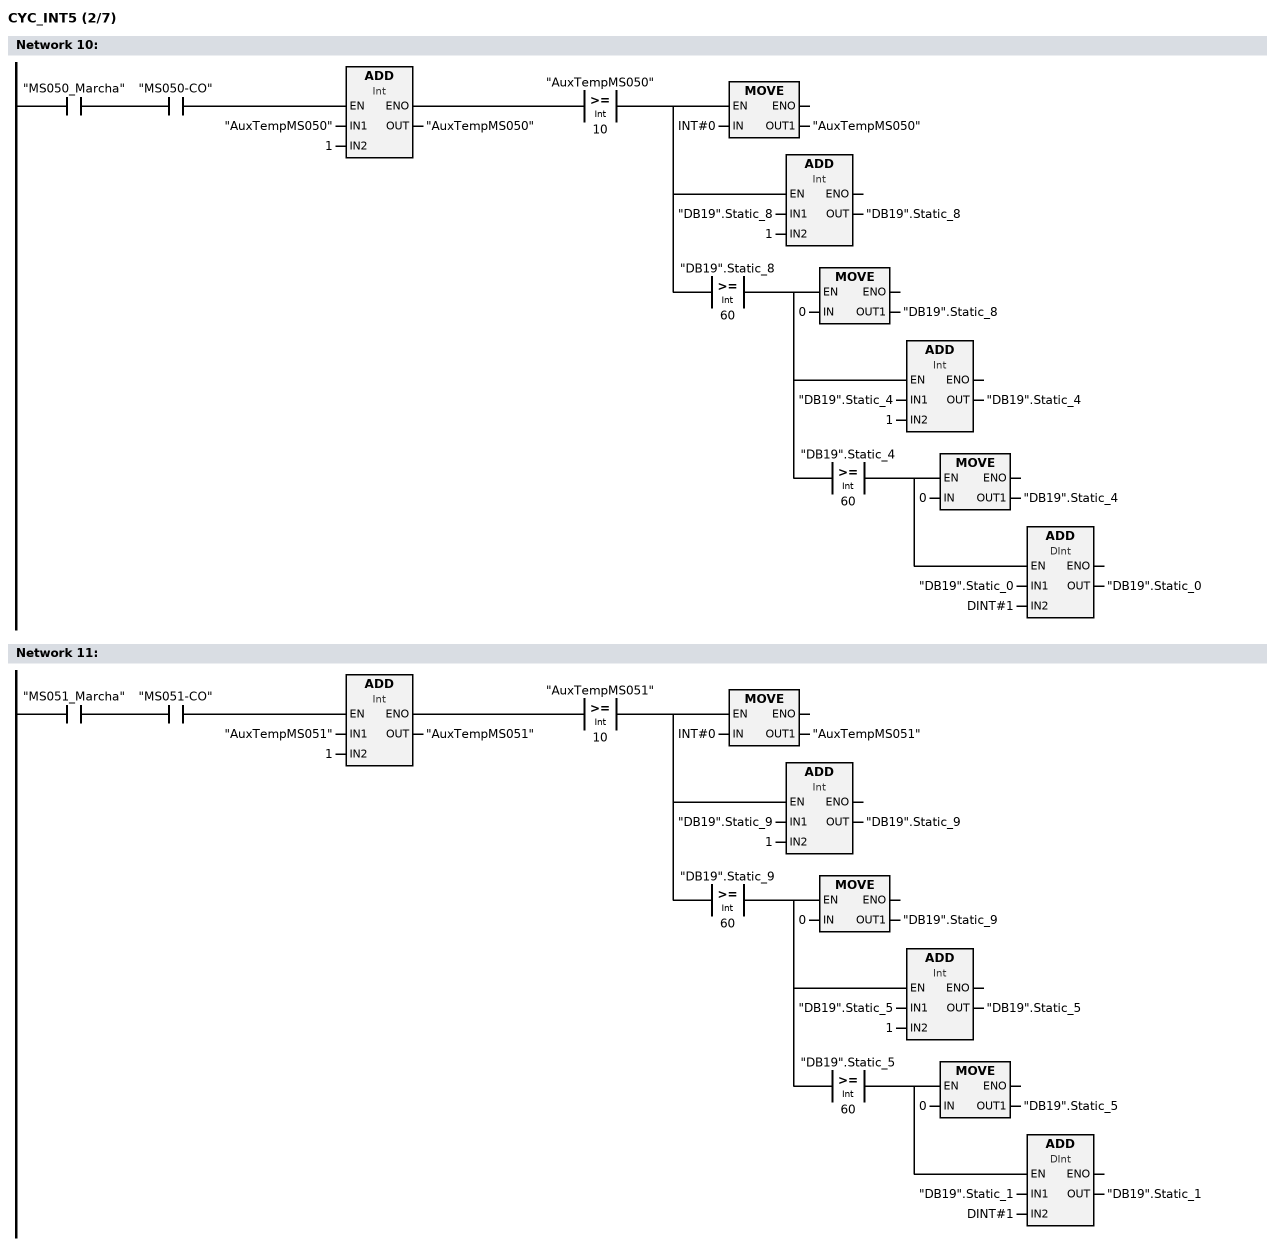
   RUNG wire#powerrail
      Contact( "MS050_Marcha" )
      Contact( "MS050-CO" )
      { S7_Templates := "SrcType := Int"; S7_GenerateENO := "TRUE" } Add(in1 := "AuxTempMS050", in2 := 1, out => "AuxTempMS050")
      { S7_Templates := "SrcType := Int" } GE_Contact(in1 := "AuxTempMS050", in2 := 10)
      wire#w1
      { S7_GenerateENO := "TRUE" } Move(in := INT#0, out1 => "AuxTempMS050")
   END_RUNG
   RUNG wire#w1
      { S7_Templates := "SrcType := Int"; S7_GenerateENO := "TRUE" } Add(in1 := "DB19".Static_8, in2 := 1, out => "DB19".Static_8)
   END_RUNG
   RUNG wire#w1
      { S7_Templates := "SrcType := Int" } GE_Contact(in1 := "DB19".Static_8, in2 := 60)
      wire#w2
      { S7_GenerateENO := "TRUE" } Move(in := 0, out1 => "DB19".Static_8)
   END_RUNG
   RUNG wire#w2
      { S7_Templates := "SrcType := Int"; S7_GenerateENO := "TRUE" } Add(in1 := "DB19".Static_4, in2 := 1, out => "DB19".Static_4)
   END_RUNG
   RUNG wire#w2
      { S7_Templates := "SrcType := Int" } GE_Contact(in1 := "DB19".Static_4, in2 := 60)
      wire#w3
      { S7_GenerateENO := "TRUE" } Move(in := 0, out1 => "DB19".Static_4)
   END_RUNG
   RUNG wire#w3
      { S7_Templates := "SrcType := DInt"; S7_GenerateENO := "TRUE" } Add(in1 := "DB19".Static_0, in2 := DINT#1, out => "DB19".Static_0)
   END_RUNG
   // the same network as SCL:
   // ENO of a box is taken as its EN; it also drops when the box reports an error
   #_w1 := "MS050_Marcha" AND "MS050-CO";
   IF #_w1 THEN "AuxTempMS050" := "AuxTempMS050" + 1; END_IF;
   #_w2 := #_w1 AND ("AuxTempMS050" >= 10);
   IF #_w2 THEN
       "AuxTempMS050" := INT#0;
       "DB19".Static_8 := "DB19".Static_8 + 1;
   END_IF;
   #_w3 := #_w2 AND ("DB19".Static_8 >= 60);
   IF #_w3 THEN
       "DB19".Static_8 := 0;
       "DB19".Static_4 := "DB19".Static_4 + 1;
   END_IF;
   #_w4 := #_w3 AND ("DB19".Static_4 >= 60);
   IF #_w4 THEN
       "DB19".Static_4 := 0;
       "DB19".Static_0 := "DB19".Static_0 + DINT#1;
   END_IF;
END_REGION

REGION Network 11
   RUNG wire#powerrail
      Contact( "MS051_Marcha" )
      Contact( "MS051-CO" )
      { S7_Templates := "SrcType := Int"; S7_GenerateENO := "TRUE" } Add(in1 := "AuxTempMS051", in2 := 1, out => "AuxTempMS051")
      { S7_Templates := "SrcType := Int" } GE_Contact(in1 := "AuxTempMS051", in2 := 10)
      wire#w1
      { S7_GenerateENO := "TRUE" } Move(in := INT#0, out1 => "AuxTempMS051")
   END_RUNG
   RUNG wire#w1
      { S7_Templates := "SrcType := Int"; S7_GenerateENO := "TRUE" } Add(in1 := "DB19".Static_9, in2 := 1, out => "DB19".Static_9)
   END_RUNG
   RUNG wire#w1
      { S7_Templates := "SrcType := Int" } GE_Contact(in1 := "DB19".Static_9, in2 := 60)
      wire#w2
      { S7_GenerateENO := "TRUE" } Move(in := 0, out1 => "DB19".Static_9)
   END_RUNG
   RUNG wire#w2
      { S7_Templates := "SrcType := Int"; S7_GenerateENO := "TRUE" } Add(in1 := "DB19".Static_5, in2 := 1, out => "DB19".Static_5)
   END_RUNG
   RUNG wire#w2
      { S7_Templates := "SrcType := Int" } GE_Contact(in1 := "DB19".Static_5, in2 := 60)
      wire#w3
      { S7_GenerateENO := "TRUE" } Move(in := 0, out1 => "DB19".Static_5)
   END_RUNG
   RUNG wire#w3
      { S7_Templates := "SrcType := DInt"; S7_GenerateENO := "TRUE" } Add(in1 := "DB19".Static_1, in2 := DINT#1, out => "DB19".Static_1)
   END_RUNG
   // the same network as SCL:
   // ENO of a box is taken as its EN; it also drops when the box reports an error
   #_w1 := "MS051_Marcha" AND "MS051-CO";
   IF #_w1 THEN "AuxTempMS051" := "AuxTempMS051" + 1; END_IF;
   #_w2 := #_w1 AND ("AuxTempMS051" >= 10);
   IF #_w2 THEN
       "AuxTempMS051" := INT#0;
       "DB19".Static_9 := "DB19".Static_9 + 1;
   END_IF;
   #_w3 := #_w2 AND ("DB19".Static_9 >= 60);
   IF #_w3 THEN
       "DB19".Static_9 := 0;
       "DB19".Static_5 := "DB19".Static_5 + 1;
   END_IF;
   #_w4 := #_w3 AND ("DB19".Static_5 >= 60);
   IF #_w4 THEN
       "DB19".Static_5 := 0;
       "DB19".Static_1 := "DB19".Static_1 + DINT#1;
   END_IF;
END_REGION

REGION Network 12
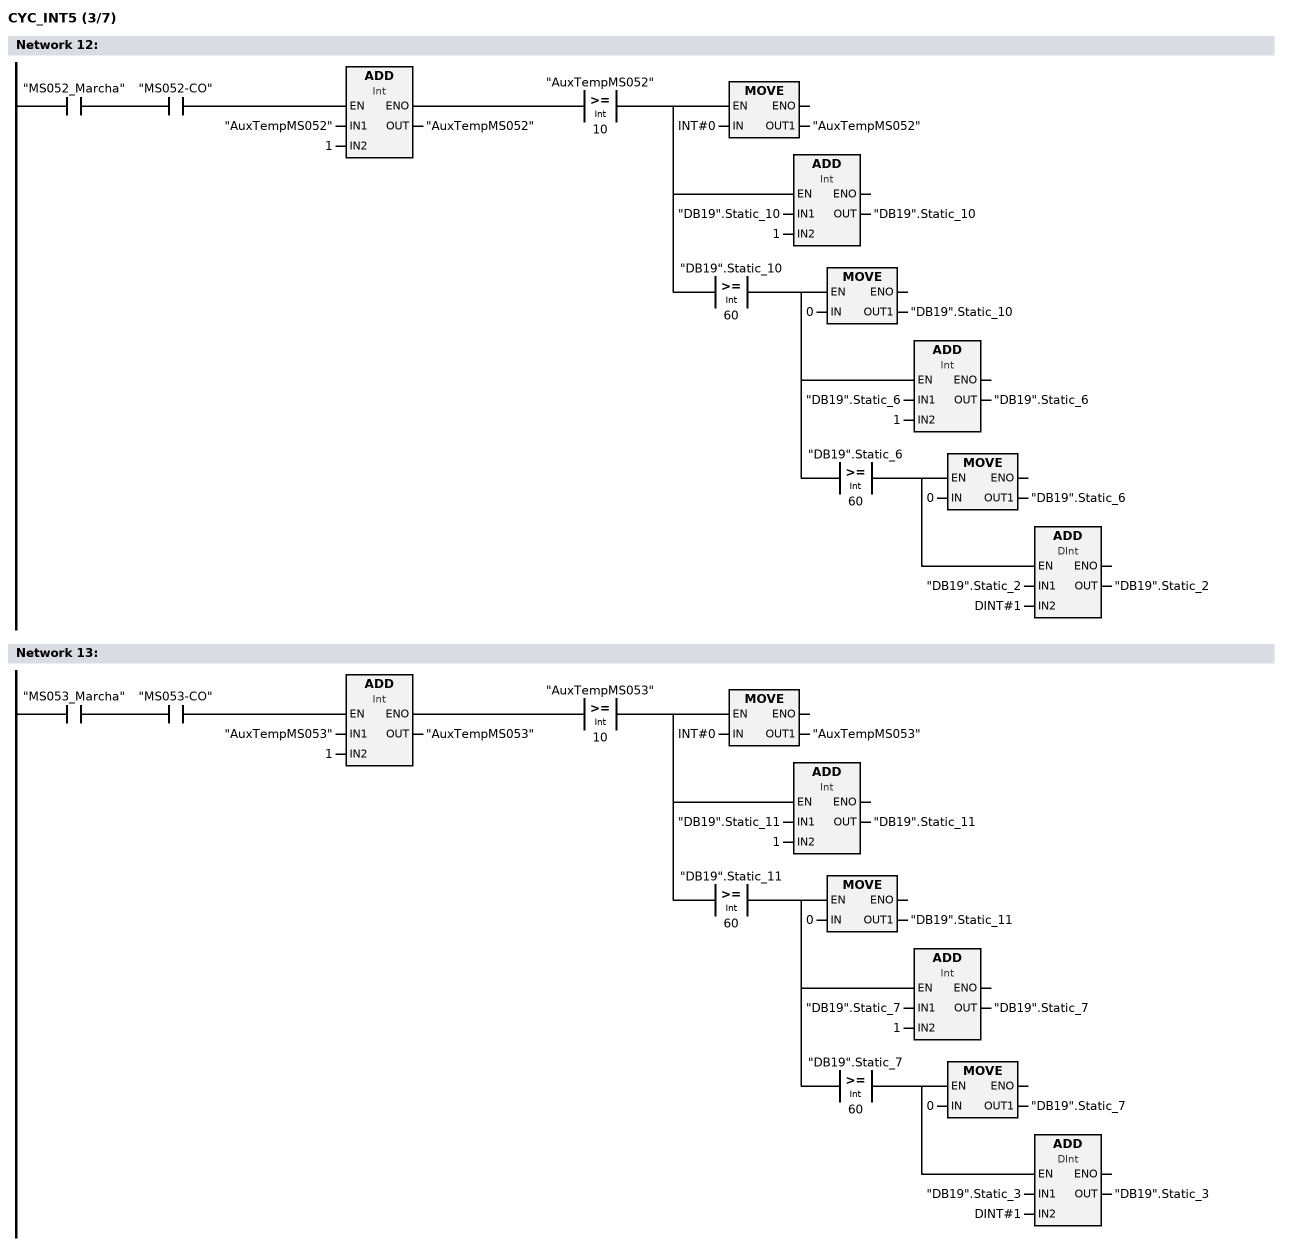
   RUNG wire#powerrail
      Contact( "MS052_Marcha" )
      Contact( "MS052-CO" )
      { S7_Templates := "SrcType := Int"; S7_GenerateENO := "TRUE" } Add(in1 := "AuxTempMS052", in2 := 1, out => "AuxTempMS052")
      { S7_Templates := "SrcType := Int" } GE_Contact(in1 := "AuxTempMS052", in2 := 10)
      wire#w1
      { S7_GenerateENO := "TRUE" } Move(in := INT#0, out1 => "AuxTempMS052")
   END_RUNG
   RUNG wire#w1
      { S7_Templates := "SrcType := Int"; S7_GenerateENO := "TRUE" } Add(in1 := "DB19".Static_10, in2 := 1, out => "DB19".Static_10)
   END_RUNG
   RUNG wire#w1
      { S7_Templates := "SrcType := Int" } GE_Contact(in1 := "DB19".Static_10, in2 := 60)
      wire#w2
      { S7_GenerateENO := "TRUE" } Move(in := 0, out1 => "DB19".Static_10)
   END_RUNG
   RUNG wire#w2
      { S7_Templates := "SrcType := Int"; S7_GenerateENO := "TRUE" } Add(in1 := "DB19".Static_6, in2 := 1, out => "DB19".Static_6)
   END_RUNG
   RUNG wire#w2
      { S7_Templates := "SrcType := Int" } GE_Contact(in1 := "DB19".Static_6, in2 := 60)
      wire#w3
      { S7_GenerateENO := "TRUE" } Move(in := 0, out1 => "DB19".Static_6)
   END_RUNG
   RUNG wire#w3
      { S7_Templates := "SrcType := DInt"; S7_GenerateENO := "TRUE" } Add(in1 := "DB19".Static_2, in2 := DINT#1, out => "DB19".Static_2)
   END_RUNG
   // the same network as SCL:
   // ENO of a box is taken as its EN; it also drops when the box reports an error
   #_w1 := "MS052_Marcha" AND "MS052-CO";
   IF #_w1 THEN "AuxTempMS052" := "AuxTempMS052" + 1; END_IF;
   #_w2 := #_w1 AND ("AuxTempMS052" >= 10);
   IF #_w2 THEN
       "AuxTempMS052" := INT#0;
       "DB19".Static_10 := "DB19".Static_10 + 1;
   END_IF;
   #_w3 := #_w2 AND ("DB19".Static_10 >= 60);
   IF #_w3 THEN
       "DB19".Static_10 := 0;
       "DB19".Static_6 := "DB19".Static_6 + 1;
   END_IF;
   #_w4 := #_w3 AND ("DB19".Static_6 >= 60);
   IF #_w4 THEN
       "DB19".Static_6 := 0;
       "DB19".Static_2 := "DB19".Static_2 + DINT#1;
   END_IF;
END_REGION

REGION Network 13
   RUNG wire#powerrail
      Contact( "MS053_Marcha" )
      Contact( "MS053-CO" )
      { S7_Templates := "SrcType := Int"; S7_GenerateENO := "TRUE" } Add(in1 := "AuxTempMS053", in2 := 1, out => "AuxTempMS053")
      { S7_Templates := "SrcType := Int" } GE_Contact(in1 := "AuxTempMS053", in2 := 10)
      wire#w1
      { S7_GenerateENO := "TRUE" } Move(in := INT#0, out1 => "AuxTempMS053")
   END_RUNG
   RUNG wire#w1
      { S7_Templates := "SrcType := Int"; S7_GenerateENO := "TRUE" } Add(in1 := "DB19".Static_11, in2 := 1, out => "DB19".Static_11)
   END_RUNG
   RUNG wire#w1
      { S7_Templates := "SrcType := Int" } GE_Contact(in1 := "DB19".Static_11, in2 := 60)
      wire#w2
      { S7_GenerateENO := "TRUE" } Move(in := 0, out1 => "DB19".Static_11)
   END_RUNG
   RUNG wire#w2
      { S7_Templates := "SrcType := Int"; S7_GenerateENO := "TRUE" } Add(in1 := "DB19".Static_7, in2 := 1, out => "DB19".Static_7)
   END_RUNG
   RUNG wire#w2
      { S7_Templates := "SrcType := Int" } GE_Contact(in1 := "DB19".Static_7, in2 := 60)
      wire#w3
      { S7_GenerateENO := "TRUE" } Move(in := 0, out1 => "DB19".Static_7)
   END_RUNG
   RUNG wire#w3
      { S7_Templates := "SrcType := DInt"; S7_GenerateENO := "TRUE" } Add(in1 := "DB19".Static_3, in2 := DINT#1, out => "DB19".Static_3)
   END_RUNG
   // the same network as SCL:
   // ENO of a box is taken as its EN; it also drops when the box reports an error
   #_w1 := "MS053_Marcha" AND "MS053-CO";
   IF #_w1 THEN "AuxTempMS053" := "AuxTempMS053" + 1; END_IF;
   #_w2 := #_w1 AND ("AuxTempMS053" >= 10);
   IF #_w2 THEN
       "AuxTempMS053" := INT#0;
       "DB19".Static_11 := "DB19".Static_11 + 1;
   END_IF;
   #_w3 := #_w2 AND ("DB19".Static_11 >= 60);
   IF #_w3 THEN
       "DB19".Static_11 := 0;
       "DB19".Static_7 := "DB19".Static_7 + 1;
   END_IF;
   #_w4 := #_w3 AND ("DB19".Static_7 >= 60);
   IF #_w4 THEN
       "DB19".Static_7 := 0;
       "DB19".Static_3 := "DB19".Static_3 + DINT#1;
   END_IF;
END_REGION

REGION Network 14
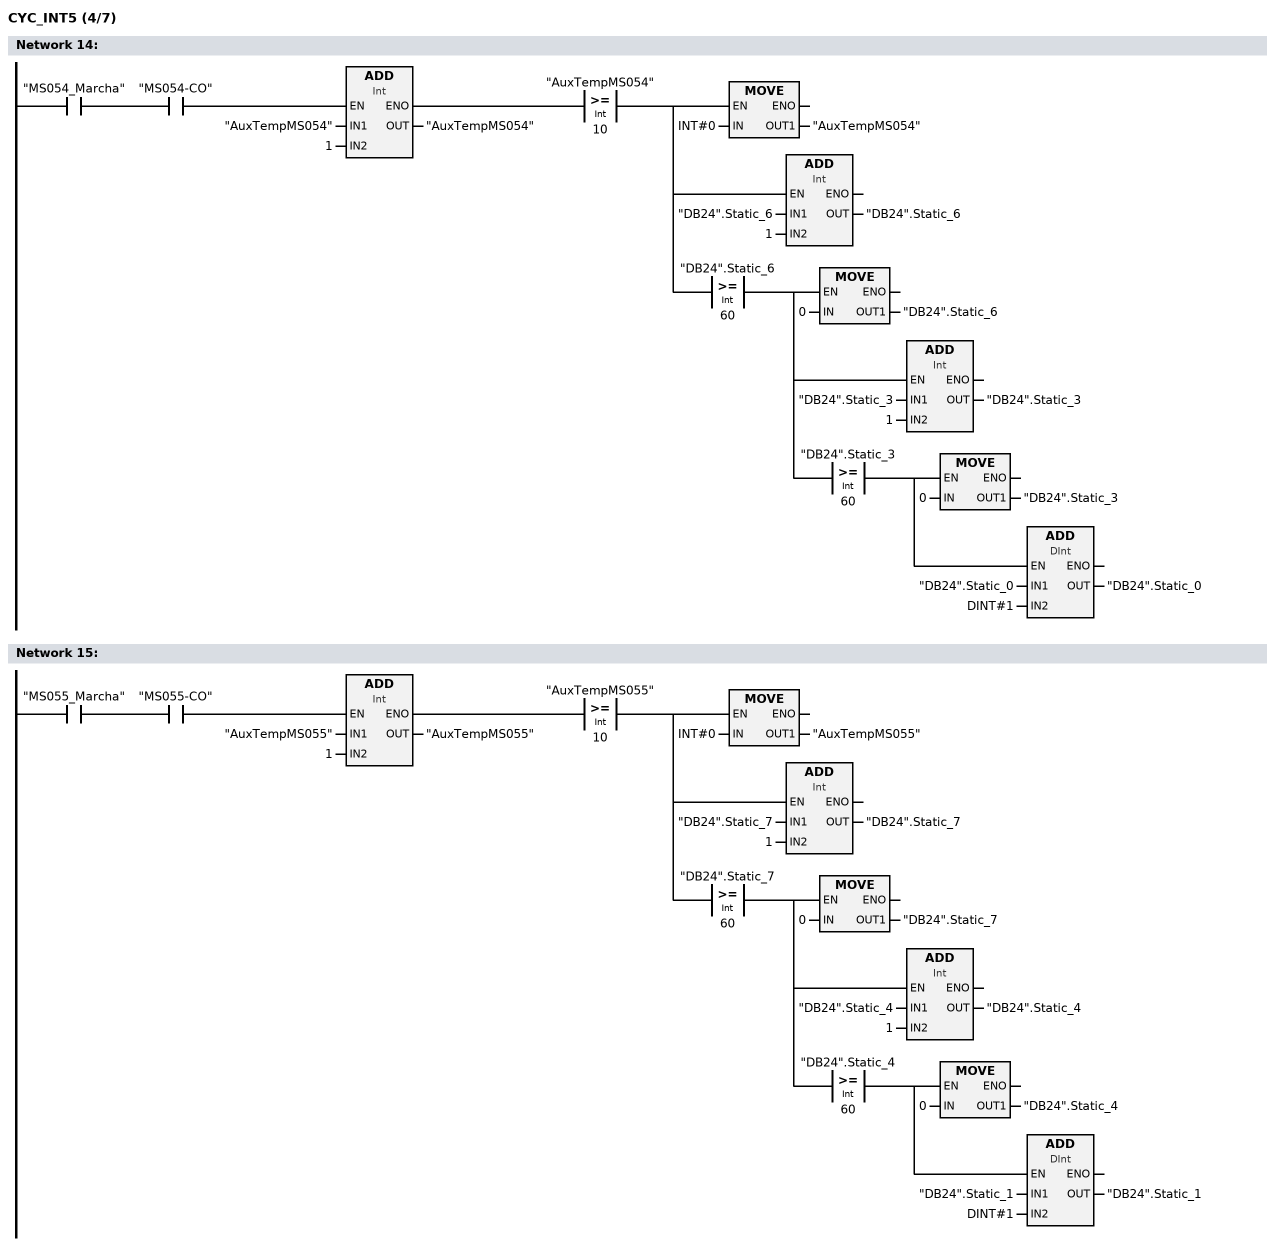
   RUNG wire#powerrail
      Contact( "MS054_Marcha" )
      Contact( "MS054-CO" )
      { S7_Templates := "SrcType := Int"; S7_GenerateENO := "TRUE" } Add(in1 := "AuxTempMS054", in2 := 1, out => "AuxTempMS054")
      { S7_Templates := "SrcType := Int" } GE_Contact(in1 := "AuxTempMS054", in2 := 10)
      wire#w1
      { S7_GenerateENO := "TRUE" } Move(in := INT#0, out1 => "AuxTempMS054")
   END_RUNG
   RUNG wire#w1
      { S7_Templates := "SrcType := Int"; S7_GenerateENO := "TRUE" } Add(in1 := "DB24".Static_6, in2 := 1, out => "DB24".Static_6)
   END_RUNG
   RUNG wire#w1
      { S7_Templates := "SrcType := Int" } GE_Contact(in1 := "DB24".Static_6, in2 := 60)
      wire#w2
      { S7_GenerateENO := "TRUE" } Move(in := 0, out1 => "DB24".Static_6)
   END_RUNG
   RUNG wire#w2
      { S7_Templates := "SrcType := Int"; S7_GenerateENO := "TRUE" } Add(in1 := "DB24".Static_3, in2 := 1, out => "DB24".Static_3)
   END_RUNG
   RUNG wire#w2
      { S7_Templates := "SrcType := Int" } GE_Contact(in1 := "DB24".Static_3, in2 := 60)
      wire#w3
      { S7_GenerateENO := "TRUE" } Move(in := 0, out1 => "DB24".Static_3)
   END_RUNG
   RUNG wire#w3
      { S7_Templates := "SrcType := DInt"; S7_GenerateENO := "TRUE" } Add(in1 := "DB24".Static_0, in2 := DINT#1, out => "DB24".Static_0)
   END_RUNG
   // the same network as SCL:
   // ENO of a box is taken as its EN; it also drops when the box reports an error
   #_w1 := "MS054_Marcha" AND "MS054-CO";
   IF #_w1 THEN "AuxTempMS054" := "AuxTempMS054" + 1; END_IF;
   #_w2 := #_w1 AND ("AuxTempMS054" >= 10);
   IF #_w2 THEN
       "AuxTempMS054" := INT#0;
       "DB24".Static_6 := "DB24".Static_6 + 1;
   END_IF;
   #_w3 := #_w2 AND ("DB24".Static_6 >= 60);
   IF #_w3 THEN
       "DB24".Static_6 := 0;
       "DB24".Static_3 := "DB24".Static_3 + 1;
   END_IF;
   #_w4 := #_w3 AND ("DB24".Static_3 >= 60);
   IF #_w4 THEN
       "DB24".Static_3 := 0;
       "DB24".Static_0 := "DB24".Static_0 + DINT#1;
   END_IF;
END_REGION

REGION Network 15
   RUNG wire#powerrail
      Contact( "MS055_Marcha" )
      Contact( "MS055-CO" )
      { S7_Templates := "SrcType := Int"; S7_GenerateENO := "TRUE" } Add(in1 := "AuxTempMS055", in2 := 1, out => "AuxTempMS055")
      { S7_Templates := "SrcType := Int" } GE_Contact(in1 := "AuxTempMS055", in2 := 10)
      wire#w1
      { S7_GenerateENO := "TRUE" } Move(in := INT#0, out1 => "AuxTempMS055")
   END_RUNG
   RUNG wire#w1
      { S7_Templates := "SrcType := Int"; S7_GenerateENO := "TRUE" } Add(in1 := "DB24".Static_7, in2 := 1, out => "DB24".Static_7)
   END_RUNG
   RUNG wire#w1
      { S7_Templates := "SrcType := Int" } GE_Contact(in1 := "DB24".Static_7, in2 := 60)
      wire#w2
      { S7_GenerateENO := "TRUE" } Move(in := 0, out1 => "DB24".Static_7)
   END_RUNG
   RUNG wire#w2
      { S7_Templates := "SrcType := Int"; S7_GenerateENO := "TRUE" } Add(in1 := "DB24".Static_4, in2 := 1, out => "DB24".Static_4)
   END_RUNG
   RUNG wire#w2
      { S7_Templates := "SrcType := Int" } GE_Contact(in1 := "DB24".Static_4, in2 := 60)
      wire#w3
      { S7_GenerateENO := "TRUE" } Move(in := 0, out1 => "DB24".Static_4)
   END_RUNG
   RUNG wire#w3
      { S7_Templates := "SrcType := DInt"; S7_GenerateENO := "TRUE" } Add(in1 := "DB24".Static_1, in2 := DINT#1, out => "DB24".Static_1)
   END_RUNG
   // the same network as SCL:
   // ENO of a box is taken as its EN; it also drops when the box reports an error
   #_w1 := "MS055_Marcha" AND "MS055-CO";
   IF #_w1 THEN "AuxTempMS055" := "AuxTempMS055" + 1; END_IF;
   #_w2 := #_w1 AND ("AuxTempMS055" >= 10);
   IF #_w2 THEN
       "AuxTempMS055" := INT#0;
       "DB24".Static_7 := "DB24".Static_7 + 1;
   END_IF;
   #_w3 := #_w2 AND ("DB24".Static_7 >= 60);
   IF #_w3 THEN
       "DB24".Static_7 := 0;
       "DB24".Static_4 := "DB24".Static_4 + 1;
   END_IF;
   #_w4 := #_w3 AND ("DB24".Static_4 >= 60);
   IF #_w4 THEN
       "DB24".Static_4 := 0;
       "DB24".Static_1 := "DB24".Static_1 + DINT#1;
   END_IF;
END_REGION

REGION Network 16
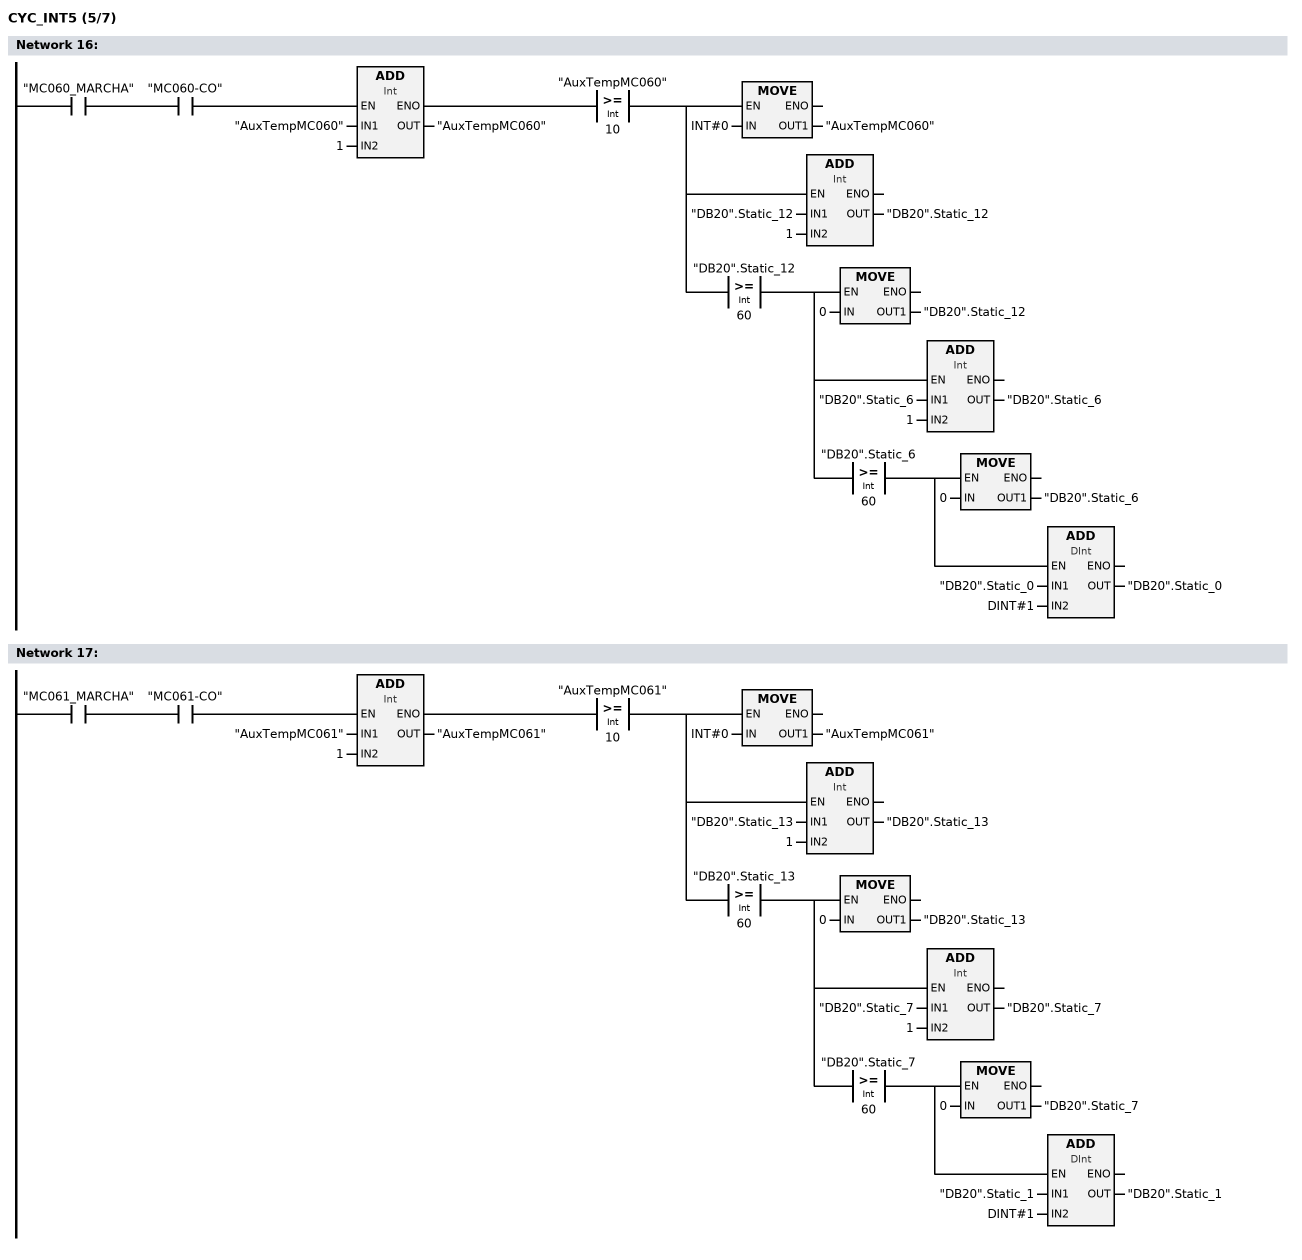
   RUNG wire#powerrail
      Contact( "MC060_MARCHA" )
      Contact( "MC060-CO" )
      { S7_Templates := "SrcType := Int"; S7_GenerateENO := "TRUE" } Add(in1 := "AuxTempMC060", in2 := 1, out => "AuxTempMC060")
      { S7_Templates := "SrcType := Int" } GE_Contact(in1 := "AuxTempMC060", in2 := 10)
      wire#w1
      { S7_GenerateENO := "TRUE" } Move(in := INT#0, out1 => "AuxTempMC060")
   END_RUNG
   RUNG wire#w1
      { S7_Templates := "SrcType := Int"; S7_GenerateENO := "TRUE" } Add(in1 := "DB20".Static_12, in2 := 1, out => "DB20".Static_12)
   END_RUNG
   RUNG wire#w1
      { S7_Templates := "SrcType := Int" } GE_Contact(in1 := "DB20".Static_12, in2 := 60)
      wire#w2
      { S7_GenerateENO := "TRUE" } Move(in := 0, out1 => "DB20".Static_12)
   END_RUNG
   RUNG wire#w2
      { S7_Templates := "SrcType := Int"; S7_GenerateENO := "TRUE" } Add(in1 := "DB20".Static_6, in2 := 1, out => "DB20".Static_6)
   END_RUNG
   RUNG wire#w2
      { S7_Templates := "SrcType := Int" } GE_Contact(in1 := "DB20".Static_6, in2 := 60)
      wire#w3
      { S7_GenerateENO := "TRUE" } Move(in := 0, out1 => "DB20".Static_6)
   END_RUNG
   RUNG wire#w3
      { S7_Templates := "SrcType := DInt"; S7_GenerateENO := "TRUE" } Add(in1 := "DB20".Static_0, in2 := DINT#1, out => "DB20".Static_0)
   END_RUNG
   // the same network as SCL:
   // ENO of a box is taken as its EN; it also drops when the box reports an error
   #_w1 := "MC060_MARCHA" AND "MC060-CO";
   IF #_w1 THEN "AuxTempMC060" := "AuxTempMC060" + 1; END_IF;
   #_w2 := #_w1 AND ("AuxTempMC060" >= 10);
   IF #_w2 THEN
       "AuxTempMC060" := INT#0;
       "DB20".Static_12 := "DB20".Static_12 + 1;
   END_IF;
   #_w3 := #_w2 AND ("DB20".Static_12 >= 60);
   IF #_w3 THEN
       "DB20".Static_12 := 0;
       "DB20".Static_6 := "DB20".Static_6 + 1;
   END_IF;
   #_w4 := #_w3 AND ("DB20".Static_6 >= 60);
   IF #_w4 THEN
       "DB20".Static_6 := 0;
       "DB20".Static_0 := "DB20".Static_0 + DINT#1;
   END_IF;
END_REGION

REGION Network 17
   RUNG wire#powerrail
      Contact( "MC061_MARCHA" )
      Contact( "MC061-CO" )
      { S7_Templates := "SrcType := Int"; S7_GenerateENO := "TRUE" } Add(in1 := "AuxTempMC061", in2 := 1, out => "AuxTempMC061")
      { S7_Templates := "SrcType := Int" } GE_Contact(in1 := "AuxTempMC061", in2 := 10)
      wire#w1
      { S7_GenerateENO := "TRUE" } Move(in := INT#0, out1 => "AuxTempMC061")
   END_RUNG
   RUNG wire#w1
      { S7_Templates := "SrcType := Int"; S7_GenerateENO := "TRUE" } Add(in1 := "DB20".Static_13, in2 := 1, out => "DB20".Static_13)
   END_RUNG
   RUNG wire#w1
      { S7_Templates := "SrcType := Int" } GE_Contact(in1 := "DB20".Static_13, in2 := 60)
      wire#w2
      { S7_GenerateENO := "TRUE" } Move(in := 0, out1 => "DB20".Static_13)
   END_RUNG
   RUNG wire#w2
      { S7_Templates := "SrcType := Int"; S7_GenerateENO := "TRUE" } Add(in1 := "DB20".Static_7, in2 := 1, out => "DB20".Static_7)
   END_RUNG
   RUNG wire#w2
      { S7_Templates := "SrcType := Int" } GE_Contact(in1 := "DB20".Static_7, in2 := 60)
      wire#w3
      { S7_GenerateENO := "TRUE" } Move(in := 0, out1 => "DB20".Static_7)
   END_RUNG
   RUNG wire#w3
      { S7_Templates := "SrcType := DInt"; S7_GenerateENO := "TRUE" } Add(in1 := "DB20".Static_1, in2 := DINT#1, out => "DB20".Static_1)
   END_RUNG
   // the same network as SCL:
   // ENO of a box is taken as its EN; it also drops when the box reports an error
   #_w1 := "MC061_MARCHA" AND "MC061-CO";
   IF #_w1 THEN "AuxTempMC061" := "AuxTempMC061" + 1; END_IF;
   #_w2 := #_w1 AND ("AuxTempMC061" >= 10);
   IF #_w2 THEN
       "AuxTempMC061" := INT#0;
       "DB20".Static_13 := "DB20".Static_13 + 1;
   END_IF;
   #_w3 := #_w2 AND ("DB20".Static_13 >= 60);
   IF #_w3 THEN
       "DB20".Static_13 := 0;
       "DB20".Static_7 := "DB20".Static_7 + 1;
   END_IF;
   #_w4 := #_w3 AND ("DB20".Static_7 >= 60);
   IF #_w4 THEN
       "DB20".Static_7 := 0;
       "DB20".Static_1 := "DB20".Static_1 + DINT#1;
   END_IF;
END_REGION

REGION Network 18
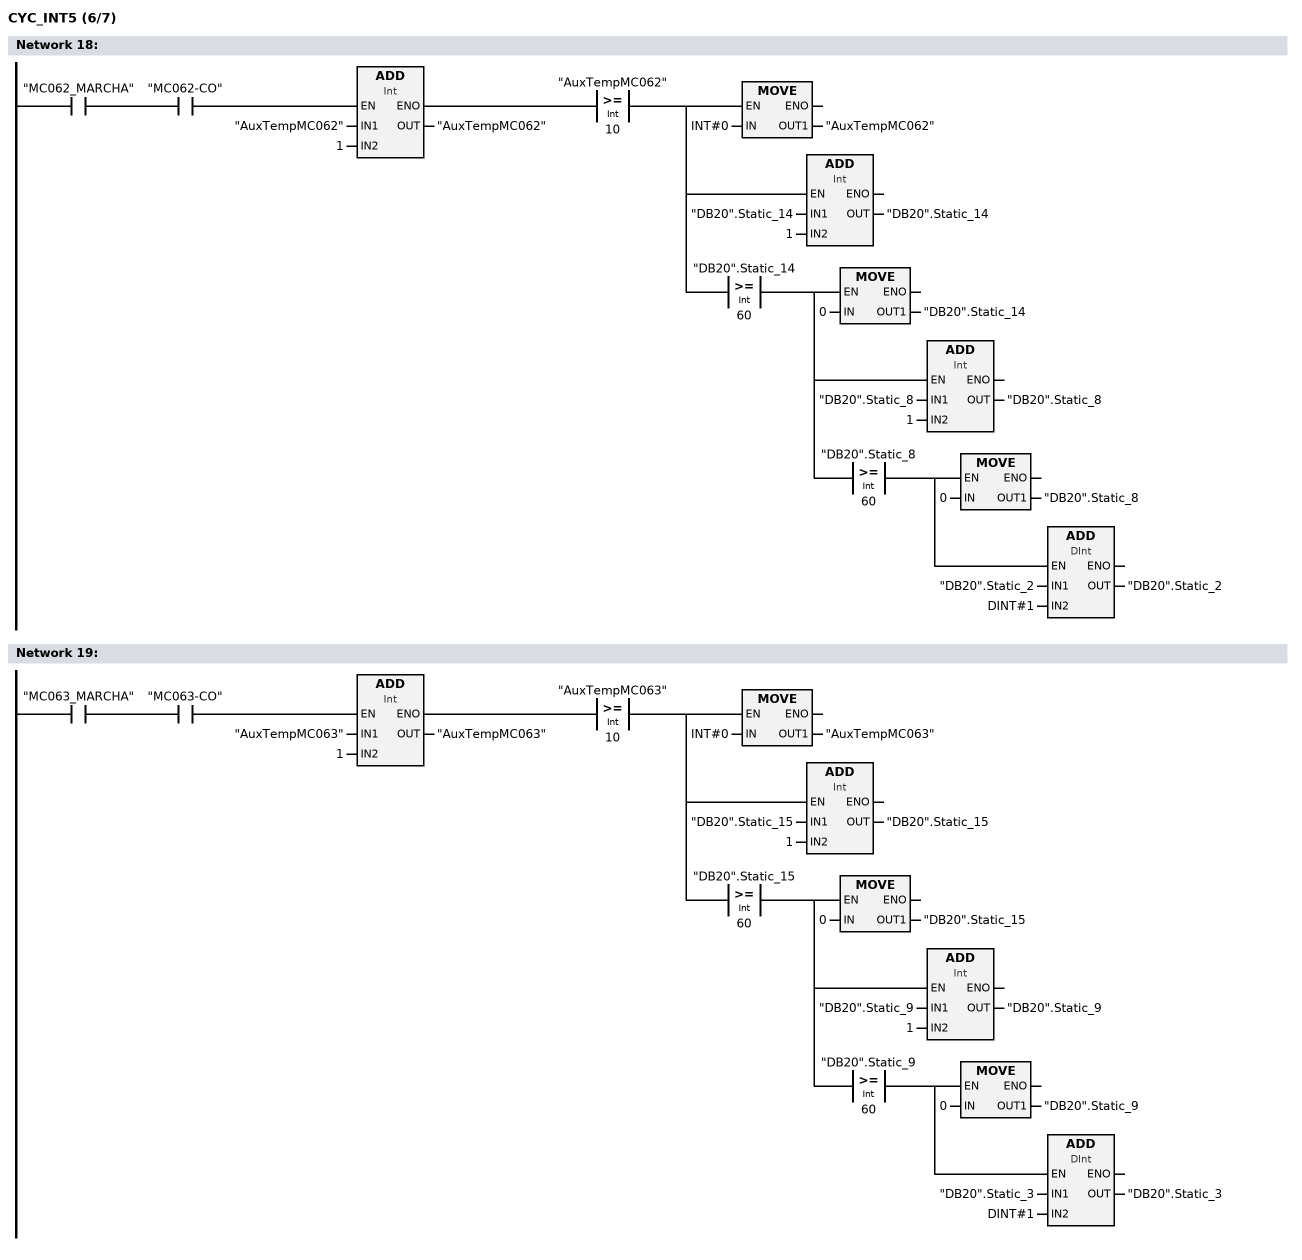
   RUNG wire#powerrail
      Contact( "MC062_MARCHA" )
      Contact( "MC062-CO" )
      { S7_Templates := "SrcType := Int"; S7_GenerateENO := "TRUE" } Add(in1 := "AuxTempMC062", in2 := 1, out => "AuxTempMC062")
      { S7_Templates := "SrcType := Int" } GE_Contact(in1 := "AuxTempMC062", in2 := 10)
      wire#w1
      { S7_GenerateENO := "TRUE" } Move(in := INT#0, out1 => "AuxTempMC062")
   END_RUNG
   RUNG wire#w1
      { S7_Templates := "SrcType := Int"; S7_GenerateENO := "TRUE" } Add(in1 := "DB20".Static_14, in2 := 1, out => "DB20".Static_14)
   END_RUNG
   RUNG wire#w1
      { S7_Templates := "SrcType := Int" } GE_Contact(in1 := "DB20".Static_14, in2 := 60)
      wire#w2
      { S7_GenerateENO := "TRUE" } Move(in := 0, out1 => "DB20".Static_14)
   END_RUNG
   RUNG wire#w2
      { S7_Templates := "SrcType := Int"; S7_GenerateENO := "TRUE" } Add(in1 := "DB20".Static_8, in2 := 1, out => "DB20".Static_8)
   END_RUNG
   RUNG wire#w2
      { S7_Templates := "SrcType := Int" } GE_Contact(in1 := "DB20".Static_8, in2 := 60)
      wire#w3
      { S7_GenerateENO := "TRUE" } Move(in := 0, out1 => "DB20".Static_8)
   END_RUNG
   RUNG wire#w3
      { S7_Templates := "SrcType := DInt"; S7_GenerateENO := "TRUE" } Add(in1 := "DB20".Static_2, in2 := DINT#1, out => "DB20".Static_2)
   END_RUNG
   // the same network as SCL:
   // ENO of a box is taken as its EN; it also drops when the box reports an error
   #_w1 := "MC062_MARCHA" AND "MC062-CO";
   IF #_w1 THEN "AuxTempMC062" := "AuxTempMC062" + 1; END_IF;
   #_w2 := #_w1 AND ("AuxTempMC062" >= 10);
   IF #_w2 THEN
       "AuxTempMC062" := INT#0;
       "DB20".Static_14 := "DB20".Static_14 + 1;
   END_IF;
   #_w3 := #_w2 AND ("DB20".Static_14 >= 60);
   IF #_w3 THEN
       "DB20".Static_14 := 0;
       "DB20".Static_8 := "DB20".Static_8 + 1;
   END_IF;
   #_w4 := #_w3 AND ("DB20".Static_8 >= 60);
   IF #_w4 THEN
       "DB20".Static_8 := 0;
       "DB20".Static_2 := "DB20".Static_2 + DINT#1;
   END_IF;
END_REGION

REGION Network 19
   RUNG wire#powerrail
      Contact( "MC063_MARCHA" )
      Contact( "MC063-CO" )
      { S7_Templates := "SrcType := Int"; S7_GenerateENO := "TRUE" } Add(in1 := "AuxTempMC063", in2 := 1, out => "AuxTempMC063")
      { S7_Templates := "SrcType := Int" } GE_Contact(in1 := "AuxTempMC063", in2 := 10)
      wire#w1
      { S7_GenerateENO := "TRUE" } Move(in := INT#0, out1 => "AuxTempMC063")
   END_RUNG
   RUNG wire#w1
      { S7_Templates := "SrcType := Int"; S7_GenerateENO := "TRUE" } Add(in1 := "DB20".Static_15, in2 := 1, out => "DB20".Static_15)
   END_RUNG
   RUNG wire#w1
      { S7_Templates := "SrcType := Int" } GE_Contact(in1 := "DB20".Static_15, in2 := 60)
      wire#w2
      { S7_GenerateENO := "TRUE" } Move(in := 0, out1 => "DB20".Static_15)
   END_RUNG
   RUNG wire#w2
      { S7_Templates := "SrcType := Int"; S7_GenerateENO := "TRUE" } Add(in1 := "DB20".Static_9, in2 := 1, out => "DB20".Static_9)
   END_RUNG
   RUNG wire#w2
      { S7_Templates := "SrcType := Int" } GE_Contact(in1 := "DB20".Static_9, in2 := 60)
      wire#w3
      { S7_GenerateENO := "TRUE" } Move(in := 0, out1 => "DB20".Static_9)
   END_RUNG
   RUNG wire#w3
      { S7_Templates := "SrcType := DInt"; S7_GenerateENO := "TRUE" } Add(in1 := "DB20".Static_3, in2 := DINT#1, out => "DB20".Static_3)
   END_RUNG
   // the same network as SCL:
   // ENO of a box is taken as its EN; it also drops when the box reports an error
   #_w1 := "MC063_MARCHA" AND "MC063-CO";
   IF #_w1 THEN "AuxTempMC063" := "AuxTempMC063" + 1; END_IF;
   #_w2 := #_w1 AND ("AuxTempMC063" >= 10);
   IF #_w2 THEN
       "AuxTempMC063" := INT#0;
       "DB20".Static_15 := "DB20".Static_15 + 1;
   END_IF;
   #_w3 := #_w2 AND ("DB20".Static_15 >= 60);
   IF #_w3 THEN
       "DB20".Static_15 := 0;
       "DB20".Static_9 := "DB20".Static_9 + 1;
   END_IF;
   #_w4 := #_w3 AND ("DB20".Static_9 >= 60);
   IF #_w4 THEN
       "DB20".Static_9 := 0;
       "DB20".Static_3 := "DB20".Static_3 + DINT#1;
   END_IF;
END_REGION

REGION Network 20
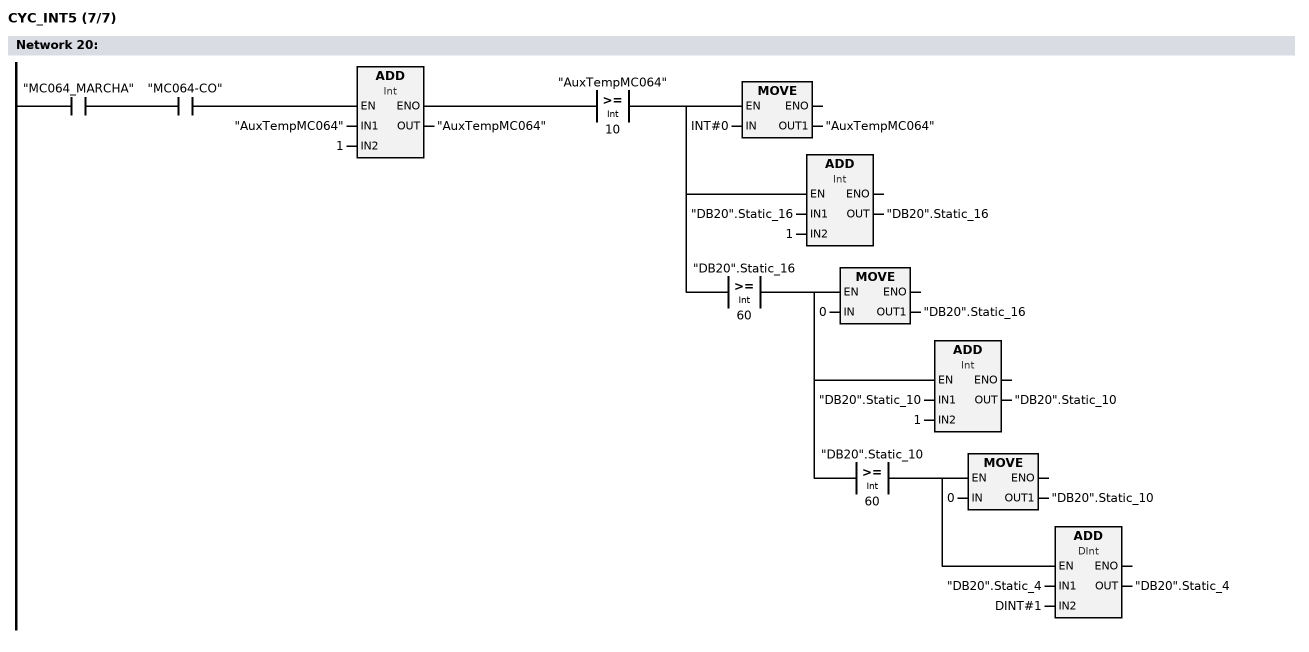
   RUNG wire#powerrail
      Contact( "MC064_MARCHA" )
      Contact( "MC064-CO" )
      { S7_Templates := "SrcType := Int"; S7_GenerateENO := "TRUE" } Add(in1 := "AuxTempMC064", in2 := 1, out => "AuxTempMC064")
      { S7_Templates := "SrcType := Int" } GE_Contact(in1 := "AuxTempMC064", in2 := 10)
      wire#w1
      { S7_GenerateENO := "TRUE" } Move(in := INT#0, out1 => "AuxTempMC064")
   END_RUNG
   RUNG wire#w1
      { S7_Templates := "SrcType := Int"; S7_GenerateENO := "TRUE" } Add(in1 := "DB20".Static_16, in2 := 1, out => "DB20".Static_16)
   END_RUNG
   RUNG wire#w1
      { S7_Templates := "SrcType := Int" } GE_Contact(in1 := "DB20".Static_16, in2 := 60)
      wire#w2
      { S7_GenerateENO := "TRUE" } Move(in := 0, out1 => "DB20".Static_16)
   END_RUNG
   RUNG wire#w2
      { S7_Templates := "SrcType := Int"; S7_GenerateENO := "TRUE" } Add(in1 := "DB20".Static_10, in2 := 1, out => "DB20".Static_10)
   END_RUNG
   RUNG wire#w2
      { S7_Templates := "SrcType := Int" } GE_Contact(in1 := "DB20".Static_10, in2 := 60)
      wire#w3
      { S7_GenerateENO := "TRUE" } Move(in := 0, out1 => "DB20".Static_10)
   END_RUNG
   RUNG wire#w3
      { S7_Templates := "SrcType := DInt"; S7_GenerateENO := "TRUE" } Add(in1 := "DB20".Static_4, in2 := DINT#1, out => "DB20".Static_4)
   END_RUNG
   // the same network as SCL:
   // ENO of a box is taken as its EN; it also drops when the box reports an error
   #_w1 := "MC064_MARCHA" AND "MC064-CO";
   IF #_w1 THEN "AuxTempMC064" := "AuxTempMC064" + 1; END_IF;
   #_w2 := #_w1 AND ("AuxTempMC064" >= 10);
   IF #_w2 THEN
       "AuxTempMC064" := INT#0;
       "DB20".Static_16 := "DB20".Static_16 + 1;
   END_IF;
   #_w3 := #_w2 AND ("DB20".Static_16 >= 60);
   IF #_w3 THEN
       "DB20".Static_16 := 0;
       "DB20".Static_10 := "DB20".Static_10 + 1;
   END_IF;
   #_w4 := #_w3 AND ("DB20".Static_10 >= 60);
   IF #_w4 THEN
       "DB20".Static_10 := 0;
       "DB20".Static_4 := "DB20".Static_4 + DINT#1;
   END_IF;
END_REGION
END_ORGANIZATION_BLOCK

// folder: Iluminación

FUNCTION "IluminaciónMTA" : Void   // FC23, LAD
{ S7_Optimized_Access := 'FALSE' }
VERSION : 0.1
   VAR_TEMP   // added for the SCL form of the ladder/FBD networks
      _s5time1 : S5Time;
   END_VAR
BEGIN

REGION Network 1
